   	Laenge_Data = SmartTags("DB_SDC_EMS_FLAGS_HEADER.LAENGE_EMS_FLAGS")
   	Allg_Offset = SmartTags("DB_SDC_EMS_FLAGS_HMI_HEADER.START_HMI")
   	HMIFlagDaten_Offset = SmartTags("DB_SDC_EMS_FLAGS_HMI_HEADER.OFFEST_HMI_DATA")
   	HMI_Nr = SmartTags("_intern_Pult_Nr")
   	
   	
      SmartTags("SDC\DB_SDC_EMS_FLAGS\_EMS_Flags_HMI_Byte_00") = 0 + HMI_Nr * (Laenge_Data + HMIFlagDaten_Offset)  - Laenge_Data - HMIFlagDaten_Offset + Allg_Offset	
      SmartTags("SDC\DB_SDC_EMS_FLAGS\_EMS_Flags_HMI_Byte_02") = 2 + HMI_Nr * (Laenge_Data + HMIFlagDaten_Offset)  - Laenge_Data - HMIFlagDaten_Offset + Allg_Offset	
      SmartTags("SDC\DB_SDC_EMS_FLAGS\_EMS_Flags_HMI_Byte_04") = 4 + HMI_Nr * (Laenge_Data + HMIFlagDaten_Offset)  - Laenge_Data - HMIFlagDaten_Offset + Allg_Offset	
      SmartTags("SDC\DB_SDC_EMS_FLAGS\_EMS_Flags_HMI_Byte_06") = 6 + HMI_Nr * (Laenge_Data + HMIFlagDaten_Offset)  - Laenge_Data - HMIFlagDaten_Offset + Allg_Offset	
      SmartTags("SDC\DB_SDC_EMS_FLAGS\_EMS_Flags_HMI_Byte_08") = 8 + HMI_Nr * (Laenge_Data + HMIFlagDaten_Offset)  - Laenge_Data - HMIFlagDaten_Offset + Allg_Offset	
      SmartTags("SDC\DB_SDC_EMS_FLAGS\_EMS_Flags_HMI_Byte_09") = 9 + HMI_Nr * (Laenge_Data + HMIFlagDaten_Offset)  - Laenge_Data - HMIFlagDaten_Offset + Allg_Offset	
      SmartTags("SDC\DB_SDC_EMS_FLAGS\_EMS_Flags_HMI_Byte_10") = 10 + HMI_Nr * (Laenge_Data + HMIFlagDaten_Offset)  - Laenge_Data - HMIFlagDaten_Offset + Allg_Offset	
      SmartTags("SDC\DB_SDC_EMS_FLAGS\_EMS_Flags_HMI_Byte_12") = 12 + HMI_Nr * (Laenge_Data + HMIFlagDaten_Offset)  - Laenge_Data - HMIFlagDaten_Offset + Allg_Offset		
      SmartTags("SDC\DB_SDC_EMS_FLAGS\_EMS_Flags_HMI_Byte_14") = 14 + HMI_Nr * (Laenge_Data + HMIFlagDaten_Offset)  - Laenge_Data - HMIFlagDaten_Offset + Allg_Offset	
      SmartTags("SDC\DB_SDC_EMS_FLAGS\_EMS_Flags_HMI_Byte_16") = 16 + HMI_Nr * (Laenge_Data + HMIFlagDaten_Offset)  - Laenge_Data - HMIFlagDaten_Offset + Allg_Offset	
      SmartTags("SDC\DB_SDC_EMS_FLAGS\_EMS_Flags_HMI_Byte_18") = 18 + HMI_Nr * (Laenge_Data + HMIFlagDaten_Offset)  - Laenge_Data - HMIFlagDaten_Offset + Allg_Offset	
      SmartTags("SDC\DB_SDC_EMS_FLAGS\_EMS_Flags_HMI_Byte_19") = 19 + HMI_Nr * (Laenge_Data + HMIFlagDaten_Offset)  - Laenge_Data - HMIFlagDaten_Offset + Allg_Offset
      SmartTags("SDC\DB_SDC_EMS_FLAGS\_EMS_Flags_HMI_Byte_20") = 20 + HMI_Nr * (Laenge_Data + HMIFlagDaten_Offset)  - Laenge_Data - HMIFlagDaten_Offset + Allg_Offset
   
      SmartTags("SDC\DB_SDC_EMS_FLAGS\DB_SDC_EMS_FLAGS.HMI[XX].EMS_Nr") = EMS_Nr
   
   '##############################################
   ' VISU sucht sich Daten:
   '##############################################

VB script "SDC_EMS_PAR"
   'HINWEIS:
   ' Beim Erstellen von Skripten können Sie mit <Strg+Leertaste> vordefinierte 
   ' Systemfunktionen in das neue Skript einbinden.
   ' Das HMIRuntime-Objekt ermöglicht einfachen Zugriff auf die Objekte des
   ' WinCC flexible Objektmodells, ihre Methoden und ihre Eigenschaften.
   ' Für ein komfortables Auswählen einer Objektreferenz betätigen Sie bitte <Alt+Rechts>.
   ' Komplexe Skripte können Sie mit Sprachelementen der Programmiersprache
   ' VBScript erstellen.
   ' Der Zugriff auf WinCC flexible Variablen erfolgt direkt über den Variablennamen,
   ' z.B. Tag = 5
   
   '________________________________________________________________________________
   '
   
   ' Groiß Andreas
   ' Siemens AG Österreich 
   ' Linz Kraußstraße 1-7 
   ' RC-AT I-IA AS-FA-SO-AE2
   ' 18.08.2015
   
   Dim EMS_Nr ' EMS Number
   Dim Laenge_Data ' Länge EMS Data
   Dim Allg_Offset ' Allg Parameter Offset
   Dim HMIParDaten_Offset ' HMI EMSdaten Offset
   
   Dim HMI_Nr ' HMI Nummer
   
   ' INIT-------------------------------------------------------------
   
   '##############################################
   ' S7 sucht sich EMSdaten:
   '##############################################
   
   Laenge_Data = SmartTags("DB_SDC_EMS_PAR_HMI_HEADER.LAENGE_PAR")
   Allg_Offset = SmartTags("DB_SDC_EMS_PAR_HMI_HEADER.START_HMI") 
   HMIParDaten_Offset = SmartTags("DB_SDC_EMS_PAR_HMI_HEADER.OFFEST_HMI_DATA")
   HMI_Nr = SmartTags("_intern_Pult_Nr")
   
   SmartTags("_PAR_HMI_Byte_00") = 0 + HMI_Nr * (Laenge_Data + HMIParDaten_Offset)  - Laenge_Data - HMIParDaten_Offset + Allg_Offset	
   SmartTags("_PAR_HMI_Byte_02") = 2 + HMI_Nr * (Laenge_Data + HMIParDaten_Offset)  - Laenge_Data - HMIParDaten_Offset + Allg_Offset	
   SmartTags("_PAR_HMI_Byte_04") = 4 + HMI_Nr * (Laenge_Data + HMIParDaten_Offset)  - Laenge_Data - HMIParDaten_Offset + Allg_Offset	
   SmartTags("_PAR_HMI_Byte_06") = 6 + HMI_Nr * (Laenge_Data + HMIParDaten_Offset)  - Laenge_Data - HMIParDaten_Offset + Allg_Offset	
   SmartTags("_PAR_HMI_Byte_08") = 8 + HMI_Nr * (Laenge_Data + HMIParDaten_Offset)  - Laenge_Data - HMIParDaten_Offset + Allg_Offset	
   SmartTags("_PAR_HMI_Byte_09") = 9 + HMI_Nr * (Laenge_Data + HMIParDaten_Offset)  - Laenge_Data - HMIParDaten_Offset + Allg_Offset
   SmartTags("_PAR_HMI_Byte_10") = 10 + HMI_Nr * (Laenge_Data + HMIParDaten_Offset)  - Laenge_Data - HMIParDaten_Offset + Allg_Offset	
   SmartTags("_PAR_HMI_Byte_12") = 12 + HMI_Nr * (Laenge_Data + HMIParDaten_Offset)  - Laenge_Data - HMIParDaten_Offset + Allg_Offset		
   SmartTags("_PAR_HMI_Byte_14") = 14 + HMI_Nr * (Laenge_Data + HMIParDaten_Offset)  - Laenge_Data - HMIParDaten_Offset + Allg_Offset	
   SmartTags("_PAR_HMI_Byte_16") = 16 + HMI_Nr * (Laenge_Data + HMIParDaten_Offset)  - Laenge_Data - HMIParDaten_Offset + Allg_Offset	
   SmartTags("_PAR_HMI_Byte_18") = 18 + HMI_Nr * (Laenge_Data + HMIParDaten_Offset)  - Laenge_Data - HMIParDaten_Offset + Allg_Offset	
   SmartTags("_PAR_HMI_Byte_19") = 19 + HMI_Nr * (Laenge_Data + HMIParDaten_Offset)  - Laenge_Data - HMIParDaten_Offset + Allg_Offset
   
   SmartTags("_Byte_EMS[XXX].DRIVE_FUNCT")  =  			0 + HMI_Nr * (Laenge_Data + HMIParDaten_Offset)  - Laenge_Data + Allg_Offset
   SmartTags("_Byte_EMS[XXX].DRIVE_V_FACT_1")  =  			2 + HMI_Nr * (Laenge_Data + HMIParDaten_Offset)  - Laenge_Data + Allg_Offset
   SmartTags("_Byte_EMS[XXX].DRIVE_V_SETP_1")  =  			6 + HMI_Nr * (Laenge_Data + HMIParDaten_Offset)  - Laenge_Data + Allg_Offset
   SmartTags("_Byte_EMS[XXX].DRIVE_V_FACT_2")  =  	   	    10 + HMI_Nr * (Laenge_Data + HMIParDaten_Offset)  - Laenge_Data + Allg_Offset
   SmartTags("_Byte_EMS[XXX].DRIVE_V_SETP_2")  =  	   		14 + HMI_Nr * (Laenge_Data + HMIParDaten_Offset)  - Laenge_Data + Allg_Offset
   SmartTags("_Byte_EMS[XXX].DRIVE_V_FACT_3")  =  	   		18 + HMI_Nr * (Laenge_Data + HMIParDaten_Offset)  - Laenge_Data + Allg_Offset
   SmartTags("_Byte_EMS[XXX].DRIVE_V_SETP_3")  =  	  		22 + HMI_Nr * (Laenge_Data + HMIParDaten_Offset)  - Laenge_Data + Allg_Offset
   SmartTags("_Byte_EMS[XXX].DRIVE_V_FACT_4")  =  	  		26 + HMI_Nr * (Laenge_Data + HMIParDaten_Offset)  - Laenge_Data + Allg_Offset
   SmartTags("_Byte_EMS[XXX].DRIVE_V_SETP_4")  =  	   		30 + HMI_Nr * (Laenge_Data + HMIParDaten_Offset)  - Laenge_Data + Allg_Offset
   SmartTags("_Byte_EMS[XXX].DRIVE_V_LIMIT_FACT")  =  		34 + HMI_Nr * (Laenge_Data + HMIParDaten_Offset)  - Laenge_Data + Allg_Offset
   SmartTags("_Byte_EMS[XXX].DRIVE_V_FACT_5")  =  	   		38 + HMI_Nr * (Laenge_Data + HMIParDaten_Offset)  - Laenge_Data + Allg_Offset
   SmartTags("_Byte_EMS[XXX].DRIVE_V_min")  =  	   		50 + HMI_Nr * (Laenge_Data + HMIParDaten_Offset)  - Laenge_Data + Allg_Offset
   SmartTags("_Byte_EMS[XXX].DRIVE_V_max_top")  =     		54 + HMI_Nr * (Laenge_Data + HMIParDaten_Offset)  - Laenge_Data + Allg_Offset
   SmartTags("_Byte_EMS[XXX].DRIVE_V_max_Not_top")  = 		58 + HMI_Nr * (Laenge_Data + HMIParDaten_Offset)  - Laenge_Data + Allg_Offset
   SmartTags("_Byte_EMS[XXX].DRIVE_V_Pos_2")  = 	   		66 + HMI_Nr * (Laenge_Data + HMIParDaten_Offset)  - Laenge_Data + Allg_Offset
   SmartTags("_Byte_EMS[XXX].DRIVE_V_Fixed_1")  = 	   		74 + HMI_Nr * (Laenge_Data + HMIParDaten_Offset)  - Laenge_Data + Allg_Offset
   SmartTags("_Byte_EMS[XXX].DRIVE_V_Fixed_2")  = 	   		78 + HMI_Nr * (Laenge_Data + HMIParDaten_Offset)  - Laenge_Data + Allg_Offset
   SmartTags("_Byte_EMS[XXX].DRIVE_V_Fixed_4_SLS_SPEED") = 86 + HMI_Nr * (Laenge_Data + HMIParDaten_Offset)  - Laenge_Data + Allg_Offset
   SmartTags("_Byte_EMS[XXX].DRIVE_V_DIV_FAST") = 			90 + HMI_Nr * (Laenge_Data + HMIParDaten_Offset)  - Laenge_Data + Allg_Offset
   SmartTags("_Byte_EMS[XXX].DRIVE_DIV_POS_FAST") = 		94 + HMI_Nr * (Laenge_Data + HMIParDaten_Offset)  - Laenge_Data + Allg_Offset
   SmartTags("_Byte_EMS[XXX].DRIVE_DIV_POS_SLOW") = 		98 + HMI_Nr * (Laenge_Data + HMIParDaten_Offset)  - Laenge_Data + Allg_Offset
   SmartTags("_Byte_EMS[XXX].DRIVE_TOL_SET_POS") = 		102 + HMI_Nr * (Laenge_Data + HMIParDaten_Offset)  - Laenge_Data + Allg_Offset
   SmartTags("_Byte_EMS[XXX].DRIVE_TOL_RESET_POS") = 		104 + HMI_Nr * (Laenge_Data + HMIParDaten_Offset)  - Laenge_Data + Allg_Offset
   SmartTags("_Byte_EMS[XXX].DRIVE_Window_Pos") = 		    106 + HMI_Nr * (Laenge_Data + HMIParDaten_Offset)  - Laenge_Data + Allg_Offset
   SmartTags("_Byte_EMS[XXX].DRIVE_Window_Overrun") = 		108 + HMI_Nr * (Laenge_Data + HMIParDaten_Offset)  - Laenge_Data + Allg_Offset
   SmartTags("_Byte_EMS[XXX].DRIVE_Window_Pos_2") = 		110 + HMI_Nr * (Laenge_Data + HMIParDaten_Offset)  - Laenge_Data + Allg_Offset
   SmartTags("_Byte_EMS[XXX].DRIVE_Window_Movement") = 	112 + HMI_Nr * (Laenge_Data + HMIParDaten_Offset)  - Laenge_Data + Allg_Offset
   SmartTags("_Byte_EMS[XXX].DRIVE_Delay_Pos") = 			116 + HMI_Nr * (Laenge_Data + HMIParDaten_Offset)  - Laenge_Data + Allg_Offset
   SmartTags("_Byte_EMS[XXX].DRIVE_DelaySpeedContr") = 	122 + HMI_Nr * (Laenge_Data + HMIParDaten_Offset)  - Laenge_Data + Allg_Offset
   SmartTags("_Byte_EMS[XXX].DRIVE_TolSpeedContr") =    	124 + HMI_Nr * (Laenge_Data + HMIParDaten_Offset)  - Laenge_Data + Allg_Offset
   
   SmartTags("_Byte_EMS[XXX].HOIST_V_min")  =  	   		140 + HMI_Nr * (Laenge_Data + HMIParDaten_Offset)  - Laenge_Data + Allg_Offset
   SmartTags("_Byte_EMS[XXX].HOIST_V_max")  =  	   		142 + HMI_Nr * (Laenge_Data + HMIParDaten_Offset)  - Laenge_Data + Allg_Offset
   SmartTags("_Byte_EMS[XXX].HOIST_V_MaxOccLift")  =  	    144 + HMI_Nr * (Laenge_Data + HMIParDaten_Offset)  - Laenge_Data + Allg_Offset
   SmartTags("_Byte_EMS[XXX].HOIST_V_Pos_1")  =  	        148 + HMI_Nr * (Laenge_Data + HMIParDaten_Offset)  - Laenge_Data + Allg_Offset
   SmartTags("_Byte_EMS[XXX].HOIST_V_Pos_2")  =  	        150 + HMI_Nr * (Laenge_Data + HMIParDaten_Offset)  - Laenge_Data + Allg_Offset
   SmartTags("_Byte_EMS[XXX].HOIST_V_Fixed_1")  =  	    152 + HMI_Nr * (Laenge_Data + HMIParDaten_Offset)  - Laenge_Data + Allg_Offset
   SmartTags("_Byte_EMS[XXX].HOIST_V_Fixed_2")  =  	    154 + HMI_Nr * (Laenge_Data + HMIParDaten_Offset)  - Laenge_Data + Allg_Offset
   SmartTags("_Byte_EMS[XXX].HOIST_V_Fixed_3")  =  	    156 + HMI_Nr * (Laenge_Data + HMIParDaten_Offset)  - Laenge_Data + Allg_Offset
   SmartTags("_Byte_EMS[XXX].HOIST_V_Fixed_4")  =  	    158 + HMI_Nr * (Laenge_Data + HMIParDaten_Offset)  - Laenge_Data + Allg_Offset
   SmartTags("_Byte_EMS[XXX].HOIST_V_Fixed_6")  =  	    162 + HMI_Nr * (Laenge_Data + HMIParDaten_Offset)  - Laenge_Data + Allg_Offset
   SmartTags("_Byte_EMS[XXX].HOIST_V_FACT_Hz_UP")  =  	    164 + HMI_Nr * (Laenge_Data + HMIParDaten_Offset)  - Laenge_Data + Allg_Offset
   SmartTags("_Byte_EMS[XXX].HOIST_V_FACT_Hz_DOWN")  =  	168 + HMI_Nr * (Laenge_Data + HMIParDaten_Offset)  - Laenge_Data + Allg_Offset
   SmartTags("_Byte_EMS[XXX].HOIST_H_Window_POS_V1")  =  	172 + HMI_Nr * (Laenge_Data + HMIParDaten_Offset)  - Laenge_Data + Allg_Offset
   SmartTags("_Byte_EMS[XXX].HOIST_H_Window_POS_V2")  =  	174 + HMI_Nr * (Laenge_Data + HMIParDaten_Offset)  - Laenge_Data + Allg_Offset
   SmartTags("_Byte_EMS[XXX].HOIST_H_TOL_SET_POS")  =  	176 + HMI_Nr * (Laenge_Data + HMIParDaten_Offset)  - Laenge_Data + Allg_Offset
   SmartTags("_Byte_EMS[XXX].HOIST_H_TOL_RESET_POS")  =  	178 + HMI_Nr * (Laenge_Data + HMIParDaten_Offset)  - Laenge_Data + Allg_Offset
   SmartTags("_Byte_EMS[XXX].HOIST_H_MIN")  =  			180 + HMI_Nr * (Laenge_Data + HMIParDaten_Offset)  - Laenge_Data + Allg_Offset
   SmartTags("_Byte_EMS[XXX].HOIST_H_MIN_without_bypass")= 182 + HMI_Nr * (Laenge_Data + HMIParDaten_Offset)  - Laenge_Data + Allg_Offset
   SmartTags("_Byte_EMS[XXX].HOIST_H_REF_OFFSET")  =  		184 + HMI_Nr * (Laenge_Data + HMIParDaten_Offset)  - Laenge_Data + Allg_Offset
   SmartTags("_Byte_EMS[XXX].HOIST_H_REF")  =  			186 + HMI_Nr * (Laenge_Data + HMIParDaten_Offset)  - Laenge_Data + Allg_Offset
   SmartTags("_Byte_EMS[XXX].HOIST_H_FACT_ENC1")  =  		188 + HMI_Nr * (Laenge_Data + HMIParDaten_Offset)  - Laenge_Data + Allg_Offset
   SmartTags("_Byte_EMS[XXX].HOIST_H_FACT_ENC2")  =  		192 + HMI_Nr * (Laenge_Data + HMIParDaten_Offset)  - Laenge_Data + Allg_Offset
   SmartTags("_Byte_EMS[XXX].HOIST_H_FACT_SPEED")  =  		196 + HMI_Nr * (Laenge_Data + HMIParDaten_Offset)  - Laenge_Data + Allg_Offset
   SmartTags("_Byte_EMS[XXX].HOIST_H_ENC_MAX_DIFF")  =  	200 + HMI_Nr * (Laenge_Data + HMIParDaten_Offset)  - Laenge_Data + Allg_Offset
   SmartTags("_Byte_EMS[XXX].HOIST_H_Slow")  =  			202 + HMI_Nr * (Laenge_Data + HMIParDaten_Offset)  - Laenge_Data + Allg_Offset
   SmartTags("_Byte_EMS[XXX].HOIST_H_tIN_POS")  =  		204 + HMI_Nr * (Laenge_Data + HMIParDaten_Offset)  - Laenge_Data + Allg_Offset
   SmartTags("_Byte_EMS[XXX].HOIST_H_REF_HMI")  =  		206 + HMI_Nr * (Laenge_Data + HMIParDaten_Offset)  - Laenge_Data + Allg_Offset

VB script "SDC_EMS_STATUS"
   'HINWEIS:
   ' Beim Erstellen von Skripten können Sie mit <Strg+Leertaste> vordefinierte 
   ' Systemfunktionen in das neue Skript einbinden.
   ' Das HMIRuntime-Objekt ermöglicht einfachen Zugriff auf die Objekte des
   ' WinCC flexible Objektmodells, ihre Methoden und ihre Eigenschaften.
   ' Für ein komfortables Auswählen einer Objektreferenz betätigen Sie bitte <Alt+Rechts>.
   ' Komplexe Skripte können Sie mit Sprachelementen der Programmiersprache
   ' VBScript erstellen.
   ' Der Zugriff auf WinCC flexible Variablen erfolgt direkt über den Variablennamen,
   ' z.B. Tag = 5
   
   '________________________________________________________________________________
   '
   
   ' Groiß Andreas
   ' Siemens AG Österreich 
   ' Linz Kraußstraße 1-7 
   ' RC-AT I-IA AS-FA-SO-AE2
   ' 23.09.2013
   
   Dim EMS_Nr ' EMS Number
   Dim Laenge_Data ' Länge EMS Data
   Dim Allg_Offset ' Allg Parameter Offset
   Dim HMIEMSDaten_Offset ' HMI EMSdaten Offset
   Dim Profil_Offset ' Allg Parameter Offset
   Dim HMI_Nr ' HMI Nummer
   
   ' INIT-------------------------------------------------------------
   SmartTags("SDC\DB_SDC_EMS\_Intern_DB_EMS_Nr") = SmartTags("DB_SDC_EMS_HMI_HEADER.DB_NR")
   
   EMS_Nr = EMS_Nr_IN
   
   If (EMS_Nr_IN < SmartTags("DB_SDC_EMS_1_HEADER.MIN_NR_EMS")) Or (EMS_Nr_IN > SmartTags("DB_SDC_EMS_1_HEADER.MAX_NR_EMS")) Then
   	EMS_Nr = SmartTags("DB_SDC_EMS_1_HEADER.MIN_NR_EMS")
   End If	
   
   If EMS_Nr_IN < 1 Then
   	EMS_Nr = 1
   End If	
   
   '##############################################
   ' S7 sucht sich EMSdaten:
   '##############################################
   
   Laenge_Data = SmartTags("DB_SDC_EMS_1_HEADER.LAENGE_EMS")
   Allg_Offset = SmartTags("DB_SDC_EMS_HMI_HEADER.START_HMI")
   HMIEMSDaten_Offset = SmartTags("DB_SDC_EMS_HMI_HEADER.OFFEST_HMI_DATA")
   HMI_Nr = SmartTags("_intern_Pult_Nr")
   
   SmartTags("SDC\DB_SDC_EMS\_EMS_HMI_Byte_00") = 0 + HMI_Nr * (Laenge_Data + HMIEMSDaten_Offset)  - Laenge_Data - HMIEMSDaten_Offset + Allg_Offset	
   SmartTags("SDC\DB_SDC_EMS\_EMS_HMI_Byte_02") = 2 + HMI_Nr * (Laenge_Data + HMIEMSDaten_Offset)  - Laenge_Data - HMIEMSDaten_Offset + Allg_Offset	
   SmartTags("SDC\DB_SDC_EMS\_EMS_HMI_Byte_04") = 4 + HMI_Nr * (Laenge_Data + HMIEMSDaten_Offset)  - Laenge_Data - HMIEMSDaten_Offset + Allg_Offset	
   SmartTags("SDC\DB_SDC_EMS\_EMS_HMI_Byte_06") = 6 + HMI_Nr * (Laenge_Data + HMIEMSDaten_Offset)  - Laenge_Data - HMIEMSDaten_Offset + Allg_Offset	
   SmartTags("SDC\DB_SDC_EMS\_EMS_HMI_Byte_08") = 8 + HMI_Nr * (Laenge_Data + HMIEMSDaten_Offset)  - Laenge_Data - HMIEMSDaten_Offset + Allg_Offset	
   SmartTags("SDC\DB_SDC_EMS\_EMS_HMI_Byte_09") = 9 + HMI_Nr * (Laenge_Data + HMIEMSDaten_Offset)  - Laenge_Data - HMIEMSDaten_Offset + Allg_Offset
   SmartTags("SDC\DB_SDC_EMS\_EMS_HMI_Byte_10") = 10 + HMI_Nr * (Laenge_Data + HMIEMSDaten_Offset)  - Laenge_Data - HMIEMSDaten_Offset + Allg_Offset	
   SmartTags("SDC\DB_SDC_EMS\_EMS_HMI_Byte_12") = 12 + HMI_Nr * (Laenge_Data + HMIEMSDaten_Offset)  - Laenge_Data - HMIEMSDaten_Offset + Allg_Offset		
   SmartTags("SDC\DB_SDC_EMS\_EMS_HMI_Byte_14") = 14 + HMI_Nr * (Laenge_Data + HMIEMSDaten_Offset)  - Laenge_Data - HMIEMSDaten_Offset + Allg_Offset	
   SmartTags("SDC\DB_SDC_EMS\_EMS_HMI_Byte_16") = 16 + HMI_Nr * (Laenge_Data + HMIEMSDaten_Offset)  - Laenge_Data - HMIEMSDaten_Offset + Allg_Offset	
   SmartTags("SDC\DB_SDC_EMS\_EMS_HMI_Byte_18") = 18 + HMI_Nr * (Laenge_Data + HMIEMSDaten_Offset)  - Laenge_Data - HMIEMSDaten_Offset + Allg_Offset	
   SmartTags("SDC\DB_SDC_EMS\_EMS_HMI_Byte_19") = 19 + HMI_Nr * (Laenge_Data + HMIEMSDaten_Offset)  - Laenge_Data - HMIEMSDaten_Offset + Allg_Offset
   
   SmartTags("SDC\DB_SDC_EMS\_Byte_EMS[XXX].IF_I_EMS.STAT") =  		0 + HMI_Nr * (Laenge_Data + HMIEMSDaten_Offset)  - Laenge_Data + Allg_Offset
   SmartTags("SDC\DB_SDC_EMS\_Byte_EMS[XXX].IF_I_EMS.ERROR") =			4 + HMI_Nr * (Laenge_Data + HMIEMSDaten_Offset)  - Laenge_Data + Allg_Offset
   SmartTags("SDC\DB_SDC_EMS\_Byte_EMS[XXX].IF_I_EMS.D_POS") =		  	6 + HMI_Nr * (Laenge_Data + HMIEMSDaten_Offset)  - Laenge_Data + Allg_Offset
   SmartTags("SDC\DB_SDC_EMS\_Byte_EMS[XXX].IF_I_EMS.H_POS") =	  		10 + HMI_Nr * (Laenge_Data + HMIEMSDaten_Offset)  - Laenge_Data + Allg_Offset
   ' SmartTags("SDC\DB_SDC_EMS\_Byte_EMS[XXX].IF_I_EMS.T_POS") =	  		12 + HMI_Nr * (Laenge_Data + HMIEMSDaten_Offset)  - Laenge_Data + Allg_Offset
   SmartTags("SDC\DB_SDC_EMS\_Byte_EMS[XXX].IF_I_EMS.EA1") =			22 + HMI_Nr * (Laenge_Data + HMIEMSDaten_Offset)  - Laenge_Data + Allg_Offset
   SmartTags("SDC\DB_SDC_EMS\_Byte_EMS[XXX].IF_I_EMS.EA2") =			26 + HMI_Nr * (Laenge_Data + HMIEMSDaten_Offset)  - Laenge_Data + Allg_Offset
   SmartTags("SDC\DB_SDC_EMS\_Byte_EMS[XXX].IF_I_EMS.EA3") =			30 + HMI_Nr * (Laenge_Data + HMIEMSDaten_Offset)  - Laenge_Data + Allg_Offset
   SmartTags("SDC\DB_SDC_EMS\_Byte_EMS[XXX].IF_Q_EMS.CONT") =		 	42 + HMI_Nr * (Laenge_Data + HMIEMSDaten_Offset)  - Laenge_Data + Allg_Offset
   SmartTags("SDC\DB_SDC_EMS\_Byte_EMS[XXX].IF_Q_EMS.D_SETPOS") =	 	46 + HMI_Nr * (Laenge_Data + HMIEMSDaten_Offset)  - Laenge_Data + Allg_Offset
   SmartTags("SDC\DB_SDC_EMS\_Byte_EMS[XXX].IF_Q_EMS.D_SETSPEED") =	50 + HMI_Nr * (Laenge_Data + HMIEMSDaten_Offset)  - Laenge_Data + Allg_Offset
   SmartTags("SDC\DB_SDC_EMS\_Byte_EMS[XXX].IF_Q_EMS.H_SETPOS") =	 	54 + HMI_Nr * (Laenge_Data + HMIEMSDaten_Offset)  - Laenge_Data + Allg_Offset
   SmartTags("SDC\DB_SDC_EMS\_Byte_EMS[XXX].IF_Q_EMS.H_SETSPEED") =	56 + HMI_Nr * (Laenge_Data + HMIEMSDaten_Offset)  - Laenge_Data + Allg_Offset
   ' SmartTags("SDC\DB_SDC_EMS\_Byte_EMS[XXX].IF_Q_EMS.T_SETPOS") =	   58 + HMI_Nr * (Laenge_Data + HMIEMSDaten_Offset)  - Laenge_Data + Allg_Offset
   ' SmartTags("SDC\DB_SDC_EMS\_Byte_EMS[XXX].IF_Q_EMS.T_SETSPEED") =	   60 + HMI_Nr * (Laenge_Data + HMIEMSDaten_Offset)  - Laenge_Data + Allg_Offset
   SmartTags("SDC\DB_SDC_EMS\_Byte_EMS[XXX].TS_STAT.VAL.ERROR") =		152 + HMI_Nr * (Laenge_Data + HMIEMSDaten_Offset)  - Laenge_Data + Allg_Offset
   SmartTags("SDC\DB_SDC_EMS\_Byte_EMS[XXX].TS_STAT.VAL.SEK") =		156 + HMI_Nr * (Laenge_Data + HMIEMSDaten_Offset)  - Laenge_Data + Allg_Offset
   SmartTags("SDC\DB_SDC_EMS\_Byte_EMS[XXX].TS_STAT.SERIES") =			164 + HMI_Nr * (Laenge_Data + HMIEMSDaten_Offset)  - Laenge_Data + Allg_Offset
   SmartTags("SDC\DB_SDC_EMS\_Byte_EMS[XXX].FKT_SET") =				190 + HMI_Nr * (Laenge_Data + HMIEMSDaten_Offset)  - Laenge_Data + Allg_Offset
   SmartTags("SDC\DB_SDC_EMS\_Byte_EMS[XXX].FLAGS") =					194 + HMI_Nr * (Laenge_Data + HMIEMSDaten_Offset)  - Laenge_Data + Allg_Offset
   SmartTags("SDC\DB_SDC_EMS\_Byte_EMS[XXX].FKT_INFO_REP_1") =			196 + HMI_Nr * (Laenge_Data + HMIEMSDaten_Offset)  - Laenge_Data + Allg_Offset
   SmartTags("SDC\DB_SDC_EMS\_Byte_EMS[XXX].FKT_INFO_REP_2") =			198 + HMI_Nr * (Laenge_Data + HMIEMSDaten_Offset)  - Laenge_Data + Allg_Offset
   SmartTags("SDC\DB_SDC_EMS\_Byte_EMS[XXX].PROFIL") =					200 + HMI_Nr * (Laenge_Data + HMIEMSDaten_Offset)  - Laenge_Data + Allg_Offset
   SmartTags("SDC\DB_SDC_EMS\_Byte_EMS[XXX].CYCLE_COUNTER") =			202 + HMI_Nr * (Laenge_Data + HMIEMSDaten_Offset)  - Laenge_Data + Allg_Offset
   SmartTags("SDC\DB_SDC_EMS\_Byte_EMS[XXX].PRECEDING_EMS") = 			204 + HMI_Nr * (Laenge_Data + HMIEMSDaten_Offset)  - Laenge_Data + Allg_Offset
   SmartTags("SDC\DB_SDC_EMS\_Byte_EMS[XXX].DISTANCE") =	 			206 + HMI_Nr * (Laenge_Data + HMIEMSDaten_Offset)  - Laenge_Data + Allg_Offset
   SmartTags("SDC\DB_SDC_EMS\_Byte_EMS[XXX].ABS_POS") =	 			210 + HMI_Nr * (Laenge_Data + HMIEMSDaten_Offset)  - Laenge_Data + Allg_Offset
   SmartTags("SDC\DB_SDC_EMS\_Byte_EMS[XXX].ERRORS_SDC") =		 		222 + HMI_Nr * (Laenge_Data + HMIEMSDaten_Offset)  - Laenge_Data + Allg_Offset
   SmartTags("SDC\DB_SDC_EMS\_Byte_EMS[XXX].VersNo[0]") =  		 	230 + HMI_Nr * (Laenge_Data + HMIEMSDaten_Offset)  - Laenge_Data + Allg_Offset
   SmartTags("SDC\DB_SDC_EMS\_Byte_EMS[XXX].VersNo[1]") =  		 	231 + HMI_Nr * (Laenge_Data + HMIEMSDaten_Offset)  - Laenge_Data + Allg_Offset
   
   SmartTags("SDC\DB_SDC_EMS\HMI[XX].EMS_Nr") = EMS_Nr
   
   '##############################################
   ' VISU Sucht sich EMSdaten:
   '##############################################
   'Laenge_EMS = SmartTags("SDC\DB_SDC_EMS\DB_SDC_EMS_1.HEADER.LAENGE_EMS")
   
   'Allg_Offset = SmartTags("SDC\DB_SDC_EMS\DB_SDC_EMS_1.HEADER.START_EMS")
   
   'SmartTags("SDC\DB_SDC_EMS\_Byte_EMS[XXX].E_I_EMS.STAT") =  			  0 + EMS_Nr * Laenge_EMS - Laenge_EMS + Allg_Offset
   
   'SmartTags("SDC\DB_SDC_EMS\_Byte_EMS[XXX].E_I_EMS.Drive_POS") =		  4 + EMS_Nr * Laenge_EMS - Laenge_EMS + Allg_Offset
   'SmartTags("SDC\DB_SDC_EMS\_Byte_EMS[XXX].E_I_EMS.Hoist_Height") =	  8 + EMS_Nr * Laenge_EMS - Laenge_EMS + Allg_Offset
   'SmartTags("SDC\DB_SDC_EMS\_Byte_EMS[XXX].E_I_EMS.FW_drive_FC") =	 10 + EMS_Nr * Laenge_EMS - Laenge_EMS + Allg_Offset
   'SmartTags("SDC\DB_SDC_EMS\_Byte_EMS[XXX].E_I_EMS.FW_hoist_FC") =	 12 + EMS_Nr * Laenge_EMS - Laenge_EMS + Allg_Offset
   'SmartTags("SDC\DB_SDC_EMS\_Byte_EMS[XXX].E_I_EMS.EA1") =			 14 + EMS_Nr * Laenge_EMS - Laenge_EMS + Allg_Offset
   'SmartTags("SDC\DB_SDC_EMS\_Byte_EMS[XXX].E_I_EMS.EA2") =			 18 + EMS_Nr * Laenge_EMS - Laenge_EMS + Allg_Offset
   'SmartTags("SDC\DB_SDC_EMS\_Byte_EMS[XXX].E_I_EMS.ERROR") =			 36 + EMS_Nr * Laenge_EMS - Laenge_EMS + Allg_Offset
   'SmartTags("SDC\DB_SDC_EMS\_Byte_EMS[XXX].A_Q_EMS.CONTROL") =		 42 + EMS_Nr * Laenge_EMS - Laenge_EMS + Allg_Offset
   'SmartTags("SDC\DB_SDC_EMS\_Byte_EMS[XXX].A_Q_EMS.DRIVE_SETPOS") =	 46 + EMS_Nr * Laenge_EMS - Laenge_EMS + Allg_Offset
   'SmartTags("SDC\DB_SDC_EMS\_Byte_EMS[XXX].A_Q_EMS.DRIVE_SETSPEED") =	 50 + EMS_Nr * Laenge_EMS - Laenge_EMS + Allg_Offset
   'SmartTags("SDC\DB_SDC_EMS\_Byte_EMS[XXX].A_Q_EMS.HOIST_SETPOS") =	 54 + EMS_Nr * Laenge_EMS - Laenge_EMS + Allg_Offset
   'SmartTags("SDC\DB_SDC_EMS\_Byte_EMS[XXX].A_Q_EMS.HOIST_SETSPEED") =	 56 + EMS_Nr * Laenge_EMS - Laenge_EMS + Allg_Offset
   'SmartTags("SDC\DB_SDC_EMS\_Byte_EMS[XXX].TS_STAT.VAL.SEK") =		180 + EMS_Nr * Laenge_EMS - Laenge_EMS + Allg_Offset
   'SmartTags("SDC\DB_SDC_EMS\_Byte_EMS[XXX].TS_STAT.SERIES") =			190 + EMS_Nr * Laenge_EMS - Laenge_EMS + Allg_Offset
   'SmartTags("SDC\DB_SDC_EMS\_Byte_EMS[XXX].FKT_SET") =				212 + EMS_Nr * Laenge_EMS - Laenge_EMS + Allg_Offset
   'SmartTags("SDC\DB_SDC_EMS\_Byte_EMS[XXX].FLAGS") =					214 + EMS_Nr * Laenge_EMS - Laenge_EMS + Allg_Offset
   'SmartTags("SDC\DB_SDC_EMS\_Byte_EMS[XXX].PROFIL") =					220 + EMS_Nr * Laenge_EMS - Laenge_EMS + Allg_Offset
   'SmartTags("SDC\DB_SDC_EMS\_Byte_EMS[XXX].PRECEDING_EMS") = 			224 + EMS_Nr * Laenge_EMS - Laenge_EMS + Allg_Offset
   'SmartTags("SDC\DB_SDC_EMS\_Byte_EMS[XXX].DISTANCE") =	 			226 + EMS_Nr * Laenge_EMS - Laenge_EMS + Allg_Offset
   'SmartTags("SDC\DB_SDC_EMS\_Byte_EMS[XXX].ABS_POS") =	 			230 + EMS_Nr * Laenge_EMS - Laenge_EMS + Allg_Offset
   'SmartTags("SDC\DB_SDC_EMS\_Byte_EMS[XXX].FAULTS_SDC") =		 		250 + EMS_Nr * Laenge_EMS - Laenge_EMS + Allg_Offset

VB script "SDC_EMS_TA_STATUS"
   'HINWEIS:
   ' Beim Erstellen von Skripten können Sie mit <Strg+Leertaste> vordefinierte 
   ' Systemfunktionen in das neue Skript einbinden.
   ' Das HMIRuntime-Objekt ermöglicht einfachen Zugriff auf die Objekte des
   ' WinCC flexible Objektmodells, ihre Methoden und ihre Eigenschaften.
   ' Für ein komfortables Auswählen einer Objektreferenz betätigen Sie bitte <Alt+Rechts>.
   ' Komplexe Skripte können Sie mit Sprachelementen der Programmiersprache
   ' VBScript erstellen.
   ' Der Zugriff auf WinCC flexible Variablen erfolgt direkt über den Variablennamen,
   ' z.B. Tag = 5
   
   '________________________________________________________________________________
   '
   
   ' Groiß Andreas
   ' Siemens AG Österreich 
   ' Linz Kraußstraße 1-7 
   ' RC-AT I-IA AS-FA-SO-AE2
   ' 12.06.2015
   
   Dim EMS_Nr ' EMS Number
   Dim Laenge_TA_Daten ' Länge TA Daten
   Dim Allg_Offset ' Allg Offset
   Dim AnzTAs	' Anzahl an TAs
   Dim OffsetEMS_TA_Daten ' Offset je EMS von TA Daten
   
   
   ' INIT-------------------------------------------------------------
   EMS_Nr = EMS_Nr_IN
   
   If (EMS_Nr_IN < SmartTags("DB_SDC_EMS_TA_HEADER.MIN_NR_EMS")) Or (EMS_Nr_IN > SmartTags("DB_SDC_EMS_TA_HEADER.MAX_NR_EMS")) Then
   	EMS_Nr = SmartTags("DB_SDC_EMS_TA_HEADER.MIN_NR_EMS")
   End If	
   
   If EMS_Nr_IN < 1 Then
   	EMS_Nr = 1
   End If	
   
   
   '##############################################
   ' VISU Sucht sich Sektions daten:
   '##############################################
   Laenge_TA_Daten = SmartTags("DB_SDC_EMS_TA_HEADER.LAENGE_TA_DATA")
   
   Allg_Offset = SmartTags("DB_SDC_EMS_TA_HEADER.START_EMS")
   
   AnzTAs = SmartTags("DB_SDC_EMS_TA_HEADER.ANZ_TA")
   
   OffsetEMS_TA_Daten = EMS_Nr * Laenge_TA_Daten * AnzTAs - Laenge_TA_Daten * AnzTAs + Allg_Offset
   
   SmartTags("_Byte_DB_SDC_EMS_TA.EMS[XX].TA1.PW1") =						  0 + 1*Laenge_TA_Daten - Laenge_TA_Daten + OffsetEMS_TA_Daten
   SmartTags("_Byte_DB_SDC_EMS_TA.EMS[XX].TA1.PW2") =						  2 + 1*Laenge_TA_Daten - Laenge_TA_Daten + OffsetEMS_TA_Daten
   SmartTags("_Byte_DB_SDC_EMS_TA.EMS[XX].TA1.PW3") =						  4 + 1*Laenge_TA_Daten - Laenge_TA_Daten + OffsetEMS_TA_Daten
   
   SmartTags("_Byte_DB_SDC_EMS_TA.EMS[XX].TA2.PW1") =						  0 + 2*Laenge_TA_Daten - Laenge_TA_Daten + OffsetEMS_TA_Daten
   SmartTags("_Byte_DB_SDC_EMS_TA.EMS[XX].TA2.PW2") =						  2 + 2*Laenge_TA_Daten - Laenge_TA_Daten + OffsetEMS_TA_Daten
   SmartTags("_Byte_DB_SDC_EMS_TA.EMS[XX].TA2.PW3") =						  4 + 2*Laenge_TA_Daten - Laenge_TA_Daten + OffsetEMS_TA_Daten
   
   SmartTags("_Byte_DB_SDC_EMS_TA.EMS[XX].TA3.PW1") =						  0 + 3*Laenge_TA_Daten - Laenge_TA_Daten + OffsetEMS_TA_Daten
   SmartTags("_Byte_DB_SDC_EMS_TA.EMS[XX].TA3.PW2") =						  2 + 3*Laenge_TA_Daten - Laenge_TA_Daten + OffsetEMS_TA_Daten
   SmartTags("_Byte_DB_SDC_EMS_TA.EMS[XX].TA3.PW3") =						  4 + 3*Laenge_TA_Daten - Laenge_TA_Daten + OffsetEMS_TA_Daten

VB script "SDC_ERROR_STAT"
   'HINWEIS:
   ' Beim Erstellen von Skripten können Sie mit <Strg+Leertaste> vordefinierte 
   ' Systemfunktionen in das neue Skript einbinden.
   ' Das HMIRuntime-Objekt ermöglicht einfachen Zugriff auf die Objekte des
   ' WinCC flexible Objektmodells, ihre Methoden und ihre Eigenschaften.
   ' Für ein komfortables Auswählen einer Objektreferenz betätigen Sie bitte <Alt+Rechts>.
   ' Komplexe Skripte können Sie mit Sprachelementen der Programmiersprache
   ' VBScript erstellen.
   ' Der Zugriff auf WinCC flexible Variablen erfolgt direkt über den Variablennamen,
   ' z.B. Tag = 5
   
   '________________________________________________________________________________
   '
   
   ' Groiß Andreas
   ' Siemens AG Österreich 
   ' Linz Kraußstraße 1-7 
   ' RC-AT I-IA AS-FA-SO-AE2
   ' 24.09.2013
   
   Dim Eintrag
   Dim Eintrag_0
   Dim Eintrag_1
   Dim Eintrag_2
   Dim Eintrag_3
   Dim Eintrag_4
   Dim Eintrag_5
   Dim Eintrag_6
   Dim Eintrag_7
   Dim Eintrag_8
   Dim Eintrag_9
   Dim Laenge_FAULT ' Länge FAULT
   Dim Allg_Offset ' Allg Parameter Offset
   
   ' INIT-------------------------------------------------------------
   SmartTags("SDC\DB_SDC_ERROR_STAT\_intern_DB_Fault_Stat_Nr") = SmartTags("DB_SDC_ERRORS_STAT_HEADER.DB_NR")
   
   Eintrag = Eintrag_Nr_IN
   
   If Eintrag_Nr_IN < SmartTags("DB_SDC_EMS_1_HEADER.MIN_NR_EMS") Or Eintrag_Nr_IN > SmartTags("DB_SDC_EMS_1_HEADER.MAX_NR_EMS") Then
   	Eintrag = SmartTags("DB_SDC_EMS_1_HEADER.MIN_NR_EMS")
   End If	
   
   If Eintrag_Nr_IN < 1 Then
   	Eintrag = 1
   End If	
   
   If Eintrag > (SmartTags("DB_SDC_ERRORS_STAT_HEADER.MAX_NR_FAULT_STAT") - SmartTags("DB_SDC_ERRORS_STAT_HEADER.FAULT_PRO_SEITE_HMI") + 1) Then
   	Eintrag = (SmartTags("DB_SDC_ERRORS_STAT_HEADER.MAX_NR_FAULT_STAT") - SmartTags("DB_SDC_ERRORS_STAT_HEADER.FAULT_PRO_SEITE_HMI") + 1)
   End If	
   
   SmartTags("SDC\DB_SDC_ERROR_STAT\_intern_Fault_Stat_Nr_Array")(0) = Eintrag + 0
   Eintrag_0 = Eintrag + 0
   SmartTags("SDC\DB_SDC_ERROR_STAT\_intern_Fault_Stat_Nr_Array")(1) = Eintrag + 1
   Eintrag_1 = Eintrag + 1
   SmartTags("SDC\DB_SDC_ERROR_STAT\_intern_Fault_Stat_Nr_Array")(2) = Eintrag + 2
   Eintrag_2 = Eintrag + 2
   SmartTags("SDC\DB_SDC_ERROR_STAT\_intern_Fault_Stat_Nr_Array")(3) = Eintrag + 3
   Eintrag_3 = Eintrag + 3
   SmartTags("SDC\DB_SDC_ERROR_STAT\_intern_Fault_Stat_Nr_Array")(4) = Eintrag + 4
   Eintrag_4 = Eintrag + 4
   SmartTags("SDC\DB_SDC_ERROR_STAT\_intern_Fault_Stat_Nr_Array")(5) = Eintrag + 5
   Eintrag_5 = Eintrag + 5
   SmartTags("SDC\DB_SDC_ERROR_STAT\_intern_Fault_Stat_Nr_Array")(6) = Eintrag + 6
   Eintrag_6 = Eintrag + 6
   SmartTags("SDC\DB_SDC_ERROR_STAT\_intern_Fault_Stat_Nr_Array")(7) = Eintrag + 7
   Eintrag_7 = Eintrag + 7
   SmartTags("SDC\DB_SDC_ERROR_STAT\_intern_Fault_Stat_Nr_Array")(8) = Eintrag + 8
   Eintrag_8 = Eintrag + 8
   SmartTags("SDC\DB_SDC_ERROR_STAT\_intern_Fault_Stat_Nr_Array")(9) = Eintrag + 9
   Eintrag_9 = Eintrag + 9
   
   Laenge_FAULT = SmartTags("DB_SDC_ERRORS_STAT_HEADER.LAENGE_FAULT_STAT")
   Allg_Offset = SmartTags("DB_SDC_ERRORS_STAT_HEADER.START_FAULT_STAT")
   
      	SmartTags("SDC\DB_SDC_ERROR_STAT\_Byte_DB_SDC_ERROR_STAT.F_STAT[XX1].EMS_TS_STAT_VAL.EMS_ID") =  			  0 + Eintrag_0 * Laenge_FAULT - Laenge_FAULT + Allg_Offset
     	SmartTags("SDC\DB_SDC_ERROR_STAT\_Byte_DB_SDC_ERROR_STAT.F_STAT[XX2].EMS_TS_STAT_VAL.EMS_ID") =  			  0 + Eintrag_1 * Laenge_FAULT - Laenge_FAULT + Allg_Offset
      	SmartTags("SDC\DB_SDC_ERROR_STAT\_Byte_DB_SDC_ERROR_STAT.F_STAT[XX3].EMS_TS_STAT_VAL.EMS_ID") =  			  0 + Eintrag_2 * Laenge_FAULT - Laenge_FAULT + Allg_Offset
     	SmartTags("SDC\DB_SDC_ERROR_STAT\_Byte_DB_SDC_ERROR_STAT.F_STAT[XX4].EMS_TS_STAT_VAL.EMS_ID") =  			  0 + Eintrag_3 * Laenge_FAULT - Laenge_FAULT + Allg_Offset
      	SmartTags("SDC\DB_SDC_ERROR_STAT\_Byte_DB_SDC_ERROR_STAT.F_STAT[XX5].EMS_TS_STAT_VAL.EMS_ID") =  			  0 + Eintrag_4 * Laenge_FAULT - Laenge_FAULT + Allg_Offset
     	SmartTags("SDC\DB_SDC_ERROR_STAT\_Byte_DB_SDC_ERROR_STAT.F_STAT[XX6].EMS_TS_STAT_VAL.EMS_ID") =  			  0 + Eintrag_5 * Laenge_FAULT - Laenge_FAULT + Allg_Offset
      	SmartTags("SDC\DB_SDC_ERROR_STAT\_Byte_DB_SDC_ERROR_STAT.F_STAT[XX7].EMS_TS_STAT_VAL.EMS_ID") =  			  0 + Eintrag_6 * Laenge_FAULT - Laenge_FAULT + Allg_Offset
     	SmartTags("SDC\DB_SDC_ERROR_STAT\_Byte_DB_SDC_ERROR_STAT.F_STAT[XX8].EMS_TS_STAT_VAL.EMS_ID") =  			  0 + Eintrag_7 * Laenge_FAULT - Laenge_FAULT + Allg_Offset
     	SmartTags("SDC\DB_SDC_ERROR_STAT\_Byte_DB_SDC_ERROR_STAT.F_STAT[XX9].EMS_TS_STAT_VAL.EMS_ID") =  			  0 + Eintrag_8 * Laenge_FAULT - Laenge_FAULT + Allg_Offset
     	SmartTags("SDC\DB_SDC_ERROR_STAT\_Byte_DB_SDC_ERROR_STAT.F_STAT[X10].EMS_TS_STAT_VAL.EMS_ID") =  			  0 + Eintrag_9 * Laenge_FAULT - Laenge_FAULT + Allg_Offset